(* Logix 5000 project; controller FV vendor 1 type 14 code 217 rev 31.11; software revision 31.00; part 53 of 63 *)
(* tags used below, declared in another part *)
   CWD : CHECKWORD_FLAGS;
   Dummy : BOOL;
   FV_AV1 : PlantItem;   // AV1
   FV_AV2 : PlantItem;   // AV2
   FV_AV2_CloseDelay : TIMER;
   FV_AV3 : PlantItem;   // AV3
   FV_AV4 : PlantItem;   // AV4
   FV_AV5 : PlantItem;   // AV5
   FV_B62 : INT[255];   // RESEED FLG
   FV_B62_0_2_OutputBit : BOOL;
   FV_bit_to_set : DINT;
   FV_data_file_address : INT;
   fv_data_file_value_to_move : DINT;
   FV_N110 : INT[255];   // FV DATA 0 CURRENT FV DATA
   FV_N111 : INT[50];   // FV1, CURRENT FV DATA
   FV_N112 : INT[50];   // FV2, CURRENT FV DATA
   FV_N113 : INT[50];   // FV3, CURRENT FV DATA
   FV_N114 : INT[50];   // FV4, CURRENT FV DATA
   FV_N115 : INT[50];   // FV5, CURRENT FV DATA
   FV_N116 : INT[50];   // FV6, CURRENT FV DATA
   FV_N117 : INT[50];   // FV7, CURRENT FV DATA
   FV_N118 : INT[50];   // FV8, CURRENT FV DATA
   FV_N119 : INT[50];   // FV9, CURRENT FV DATA
   FV_N12 : INT[255];   // SYS_PARMS System Parameter Fil e
   FV_N120 : INT[50];   // FV10, CURRENT FV DATA
   FV_N121 : INT[50];   // FV11, CURRENT FV DATA
   FV_N122 : INT[50];   // FV12, CURRENT FV DATA
   FV_N123 : INT[50];   // FV13, CURRENT FV DATA
   FV_N124 : INT[50];   // FV14, CURRENT FV DATA
   FV_N125 : INT[50];   // FV15, CURRENT FV DATA
   FV_N126 : INT[50];   // FV16, CURRENT FV DATA
   FV_N127 : INT[50];   // FV17, CURRENT FV DATA
   FV_N128 : INT[50];   // FV18, CURRENT FV DATA
   FV_N129 : INT[50];   // FV19, CURRENT FV DATA
   FV_N130 : INT[50];   // FV20, CURRENT FV DATA
   FV_N131 : INT[50];   // FV21, CURRENT FV DATA
   FV_N132 : INT[50];   // FV22, CURRENT FV DATA
   FV_N133 : INT[50];   // FV23, CURRENT FV DATA
   FV_N134 : INT[50];   // FV24, CURRENT FV DATA
   FV_N135 : INT[50];   // FV25, CURRENT FV DATA
   FV_N136 : INT[50];   // YSV1, CURRENT FV DATA
   FV_N137 : INT[50];   // YSV2, CURRENT FV DATA
   FV_N138 : INT[50];   // YSV3, CURRENT FV DATA
   FV_N139 : INT[255];   // YST1
   FV_N14 : INT[255];   // ME>PLC Inter PLC comms traf fic outbound
   FV_N140 : INT[255];   // YST2
   FV_N141 : INT[255];   // YSV1 DATA
   FV_N142 : INT[255];   // YSV2 DATA
   FV_N143 : INT[255];   // YSV3 DATA
   FV_N144 : INT[255];   // YST1 DATA
   FV_N145 : INT[255];   // YST2 DATA
   FV_N146 : INT[50];   // FV26, CURRENT FV DATA
   FV_N147 : INT[50];   // FV27, CURRENT FV DATA
   FV_N148 : INT[50];   // FV28, CURRENT FV DATA
   FV_N149 : INT[50];   // FV29, CURRENT FV DATA
   FV_N150 : INT[50];   // FV30, CURRENT FV DATA
   FV_N151 : INT[50];   // FV31, CURRENT FV DATA
   FV_N60 : INT[255];   // RESEED<PC
   FV_N61 : INT[255];   // RESEED>PC
   FV_N64 : INT[255];   // RESEED_SV
   FV_SOV2 : PlantItem;   // SOV2
   FV_T63 : TIMER[20];
   FV_word_offset : INT;
   FV_YSV1R : PlantItem;   // YSV1R
   Reseeding_transaction_log_delay : DINT;
(* FV_Common, continued *)

ROUTINE FV_RESEED_MC_30   (* ladder *)
   // Run Reseeding  command interpreter
   0: JSR(FV_RESEED_CP_31,0);
   // Run Reseeding Process If Active
   1: XIC(FV_B62[0].0)JSR(FV_RESEED_PRO_32,0);
   // PostScan reseeding process if not active.
   2: XIO(FV_B62[0].0)OSR(FV_B62[0].2,FV_B62_0_2_OutputBit)XIC(FV_B62_0_2_OutputBit)JSR(FV_RESEED_PRO_32,0);
END_ROUTINE

ROUTINE FV_RESEED_PRO_32   (* ladder *)
   // Yeast reseeding process control routine Step 10: Initialise
   0: XIC(FV_B62[0].1)EQU(FV_N61[1],10)MCR();
   // Set restart step for this process
   1: MOV(10,FV_N61[3]);
   // Make pointer toYSV's data file
   2: ADD(FV_N60[1],140,FV_N61[15]);
   // Make pointer to YSV's Attemporation Data File
   3: MOV(136,FV_N61[14]);
   // Make pointer to FV's attemperation data file.
   4: ADD(FV_N60[3],110,FV_N61[13]);
   // Zero PC total transferred display register.
   5: CLR(FV_N61[10]);
   // Initialise reseeding process timers.
   6: [RES(FV_T63[3]) ,RES(FV_T63[7]) ,MUL(FV_N12[10],1000,FV_T63[3].PRE) ,MUL(FV_N12[11],1000,FV_T63[4].PRE) ,MUL(FV_N12[12],1000,FV_T63[5].PRE) ];
   // Initialise reseeding process timers.
   7: OTU(FV_B62[1].0);
   // Advance to next step
   8: MOV(20,FV_N61[1]);
   9: MCR();
   // Step 20: Rouse YSV and displace water from transfer line.
   10: XIC(FV_B62[0].1)EQU(FV_N61[1],20)MCR();
   11: MOV(20,FV_N61[3]);
   12: [TON(FV_T63[4],?,?) ,XIC(FV_T63[4].DN) MOV(30,FV_N61[1]) ];
   13: MCR();
   // Step 30: Initialise transfer registers.
   14: XIC(FV_B62[0].1)EQU(FV_N61[1],30)MCR();
   // Set restart step for this process
   15: MOV(30,FV_N61[3]);
   16: TON(FV_T63[6],?,?);
   // Save YSV volume at start of transfer
   17: JSR(FV_Get_FV_Datafile_Value,2,FV_N61[15],5)MOV(fv_data_file_value_to_move,FV_N61[17]);
   // Calculate maximum allowed weight in YSV before alarm
   18: ADD(FV_N61[17],FV_N12[4],FV_N61[18]);
   // Calculate volume at which to stop discharging vessel. If < 0 , set to zero.
   19: [SUB(FV_N61[17],FV_N60[2],FV_N61[21]) ,LES(FV_N61[21],0) MOV(0,FV_N61[21]) ];
   // Advance to next step.
   20: XIC(FV_T63[6].DN)MOV(40,FV_N61[1]);
   // Advance to next step.
   21: MCR();
   // Step 40: transfer yeast to centrifuge main until target volume reached.
   22: XIC(FV_B62[0].1)EQU(FV_N61[1],40)MCR();
   23: MOV(40,FV_N61[3]);
   // Calculate total volume transferred to centrifuge main so far for PC display (zero if < 0).
   24: [JSR(FV_Get_FV_Datafile_Value,2,FV_N61[15],5) SUB(FV_N61[17],fv_data_file_value_to_move,FV_N61[10]) ,LES(FV_N61[10],0) MOV(0,FV_N61[10]) ];
   // Advance to next step if current YSV volume is less than or equal to target end volume.
   25: JSR(FV_Get_FV_Datafile_Value,2,FV_N61[15],5)LEQ(fv_data_file_value_to_move,FV_N61[21])MOV(50,FV_N61[1]);
   // Generate alarm if YSV weight increases whilst vessel is transfering
   26: JSR(FV_Get_FV_Datafile_Value,2,FV_N61[15],5)GRT(fv_data_file_value_to_move,FV_N61[18])[MOV(500,FV_N61[4]) ,MOV(FV_N60[1],FV_N61[5]) ,ADD(fv_data_file_value_to_move,FV_N12[4],FV_N61[18]) ];
   27: MCR();
   // Step 50: Flush yeast to drain with water.
   28: XIC(FV_B62[0].1)EQU(FV_N61[1],50)MCR();
   29: MOV(50,FV_N61[3]);
   // Allow time for AV4 to close before opening AV3
   30: TON(FV_T63[7],?,?);
   // Time the water flush
   31: XIC(FV_T63[7].DN)[TON(FV_T63[5],?,?) ,XIC(FV_T63[5].DN) TON(FV_AV2_CloseDelay,?,?) ,XIC(FV_AV2_CloseDelay.DN) MOV(60,FV_N61[1]) ];
   32: MCR();
   // Step 60: Save transfer data for PC and reset YSV.
   33: XIC(FV_B62[0].1)EQU(FV_N61[1],60)MCR();
   34: [MOV(FV_N60[1],FV_N64[1]) ,MOV(FV_N61[10],FV_N64[2]) ,MOV(FV_N60[3],FV_N64[3]) ,MOV(FV_N60[4],FV_N64[4]) ,OTL(FV_N64[0].0) ];
   35: MOV(1,Reseeding_transaction_log_delay);
   // Send MV number which was reseeded to MV attemporation system so it can set control to ageing
   36: [LIM(29,FV_N60[4],56) ,EQU(FV_N60[4],94) ,LIM(336,FV_N60[4],347) ][MOV(FV_N60[4],FV_N14[1]) ,OTL(FV_N14[2].0) ];
   // Send CT number which was reseeded to CT attemporation system so it can set control to conditioning
   37: LIM(57,FV_N60[4],91)[MOV(FV_N60[4],FV_N14[4]) ,OTL(FV_N14[5].0) ];
   38: [JSR(FV_Set_FV_Datafile_Value,3,0,FV_N61[15],3) ,JSR(FV_Set_FV_Datafile_Value,3,5,FV_N61[15],0) ];
   39: CLR(FV_N61[16]);
   40: MCR();
   // Drive valves, rouser & pump dependent on current process step.
   41: XIC(FV_B62[0].1)LIM(20,FV_N61[1],50)MCR();
   42: [RTO(FV_T63[3],?,?) ,XIC(FV_T63[3].TT) OTE(FV_YSV1R.DriveBits.3) ];
   43: [EQU(FV_N61[1],20) ,EQU(FV_N61[1],40) ]OTE(FV_AV1.DriveBits.5);
   44: EQU(FV_N61[1],50)XIC(FV_T63[7].DN)XIO(FV_AV2_CloseDelay.TT)OTE(FV_AV2.DriveBits.5);
   45: EQU(FV_N61[1],40)OTE(FV_AV4.DriveBits.5);
   46: [EQU(FV_N61[1],20) ,EQU(FV_N61[1],50) XIC(FV_T63[7].DN) ]OTE(FV_AV5.DriveBits.5);
   47: [EQU(FV_N61[1],20) ,EQU(FV_N61[1],40) ,EQU(FV_N61[1],50) ][TON(FV_T63[8],?,?) ,XIC(FV_T63[8].DN) OTE(FV_SOV2.DriveBits.1) ];
   48: MCR();
   // Alarms
   49: XIC(FV_B62[0].1)MCR();
   50: [XIC(FV_AV1.CW.[CWD.FAULT]) ,XIC(FV_AV2.CW.[CWD.FAULT]) ,XIC(FV_AV3.CW.[CWD.FAULT]) ,XIC(FV_AV4.CW.[CWD.FAULT]) ]OTU(FV_B62[0].1);
   51: GRT(FV_N61[4],0)OTU(FV_B62[0].1);
   52: XIO(FV_B62[0].1)[MOV(4,FV_N61[0]) ,OTU(FV_N61[2].2) ,OTL(FV_N61[2].3) ,OTL(FV_N61[2].4) ,MOV(0,FV_N61[1]) ];
   53: MCR();
END_ROUTINE

ROUTINE FV_Set_Flag_In_FV_Datafile   (* ladder *)
   // Routine to Set the value of something within the FV Data Files, Used to replace indirection originally used
   0: SBR(FV_data_file_address,FV_word_offset,FV_bit_to_set)OTE(Dummy);
   1: EQU(FV_data_file_address,110)OTL(FV_N110[FV_word_offset].[FV_bit_to_set]);
   2: EQU(FV_data_file_address,111)OTL(FV_N111[FV_word_offset].[FV_bit_to_set]);
   3: EQU(FV_data_file_address,112)OTL(FV_N112[FV_word_offset].[FV_bit_to_set]);
   4: EQU(FV_data_file_address,113)OTL(FV_N113[FV_word_offset].[FV_bit_to_set]);
   5: EQU(FV_data_file_address,114)OTL(FV_N114[FV_word_offset].[FV_bit_to_set]);
   6: EQU(FV_data_file_address,115)OTL(FV_N115[FV_word_offset].[FV_bit_to_set]);
   7: EQU(FV_data_file_address,116)OTL(FV_N116[FV_word_offset].[FV_bit_to_set]);
   8: EQU(FV_data_file_address,117)OTL(FV_N117[FV_word_offset].[FV_bit_to_set]);
   9: EQU(FV_data_file_address,118)OTL(FV_N118[FV_word_offset].[FV_bit_to_set]);
   10: EQU(FV_data_file_address,119)OTL(FV_N119[FV_word_offset].[FV_bit_to_set]);
   11: EQU(FV_data_file_address,120)OTL(FV_N120[FV_word_offset].[FV_bit_to_set]);
   12: EQU(FV_data_file_address,121)OTL(FV_N121[FV_word_offset].[FV_bit_to_set]);
   13: EQU(FV_data_file_address,122)OTL(FV_N122[FV_word_offset].[FV_bit_to_set]);
   14: EQU(FV_data_file_address,123)OTL(FV_N123[FV_word_offset].[FV_bit_to_set]);
   15: EQU(FV_data_file_address,124)OTL(FV_N124[FV_word_offset].[FV_bit_to_set]);
   16: EQU(FV_data_file_address,125)OTL(FV_N125[FV_word_offset].[FV_bit_to_set]);
   17: EQU(FV_data_file_address,126)OTL(FV_N126[FV_word_offset].[FV_bit_to_set]);
   18: EQU(FV_data_file_address,127)OTL(FV_N127[FV_word_offset].[FV_bit_to_set]);
   19: EQU(FV_data_file_address,128)OTL(FV_N128[FV_word_offset].[FV_bit_to_set]);
   20: EQU(FV_data_file_address,129)OTL(FV_N129[FV_word_offset].[FV_bit_to_set]);
   21: EQU(FV_data_file_address,130)OTL(FV_N130[FV_word_offset].[FV_bit_to_set]);
   22: EQU(FV_data_file_address,131)OTL(FV_N131[FV_word_offset].[FV_bit_to_set]);
   23: EQU(FV_data_file_address,132)OTL(FV_N132[FV_word_offset].[FV_bit_to_set]);
   24: EQU(FV_data_file_address,133)OTL(FV_N133[FV_word_offset].[FV_bit_to_set]);
   25: EQU(FV_data_file_address,134)OTL(FV_N134[FV_word_offset].[FV_bit_to_set]);
   26: EQU(FV_data_file_address,135)OTL(FV_N135[FV_word_offset].[FV_bit_to_set]);
   27: EQU(FV_data_file_address,136)OTL(FV_N136[FV_word_offset].[FV_bit_to_set]);
   28: EQU(FV_data_file_address,137)OTL(FV_N137[FV_word_offset].[FV_bit_to_set]);
   29: EQU(FV_data_file_address,138)OTL(FV_N138[FV_word_offset].[FV_bit_to_set]);
   30: EQU(FV_data_file_address,139)OTL(FV_N139[FV_word_offset].[FV_bit_to_set]);
   31: EQU(FV_data_file_address,140)OTL(FV_N140[FV_word_offset].[FV_bit_to_set]);
   32: EQU(FV_data_file_address,141)OTL(FV_N141[FV_word_offset].[FV_bit_to_set]);
   33: EQU(FV_data_file_address,142)OTL(FV_N142[FV_word_offset].[FV_bit_to_set]);
   34: EQU(FV_data_file_address,143)OTL(FV_N143[FV_word_offset].[FV_bit_to_set]);
   35: EQU(FV_data_file_address,144)OTL(FV_N144[FV_word_offset].[FV_bit_to_set]);
   36: EQU(FV_data_file_address,145)OTL(FV_N145[FV_word_offset].[FV_bit_to_set]);
   37: EQU(FV_data_file_address,146)OTL(FV_N146[FV_word_offset].[FV_bit_to_set]);
   38: EQU(FV_data_file_address,147)OTL(FV_N147[FV_word_offset].[FV_bit_to_set]);
   39: EQU(FV_data_file_address,148)OTL(FV_N148[FV_word_offset].[FV_bit_to_set]);
   40: EQU(FV_data_file_address,149)OTL(FV_N149[FV_word_offset].[FV_bit_to_set]);
   41: EQU(FV_data_file_address,150)OTL(FV_N150[FV_word_offset].[FV_bit_to_set]);
   42: EQU(FV_data_file_address,151)OTL(FV_N151[FV_word_offset].[FV_bit_to_set]);
   43: RET();
END_ROUTINE
